// TIA Portal project "Factory_Project_V17" (V17) (continued)
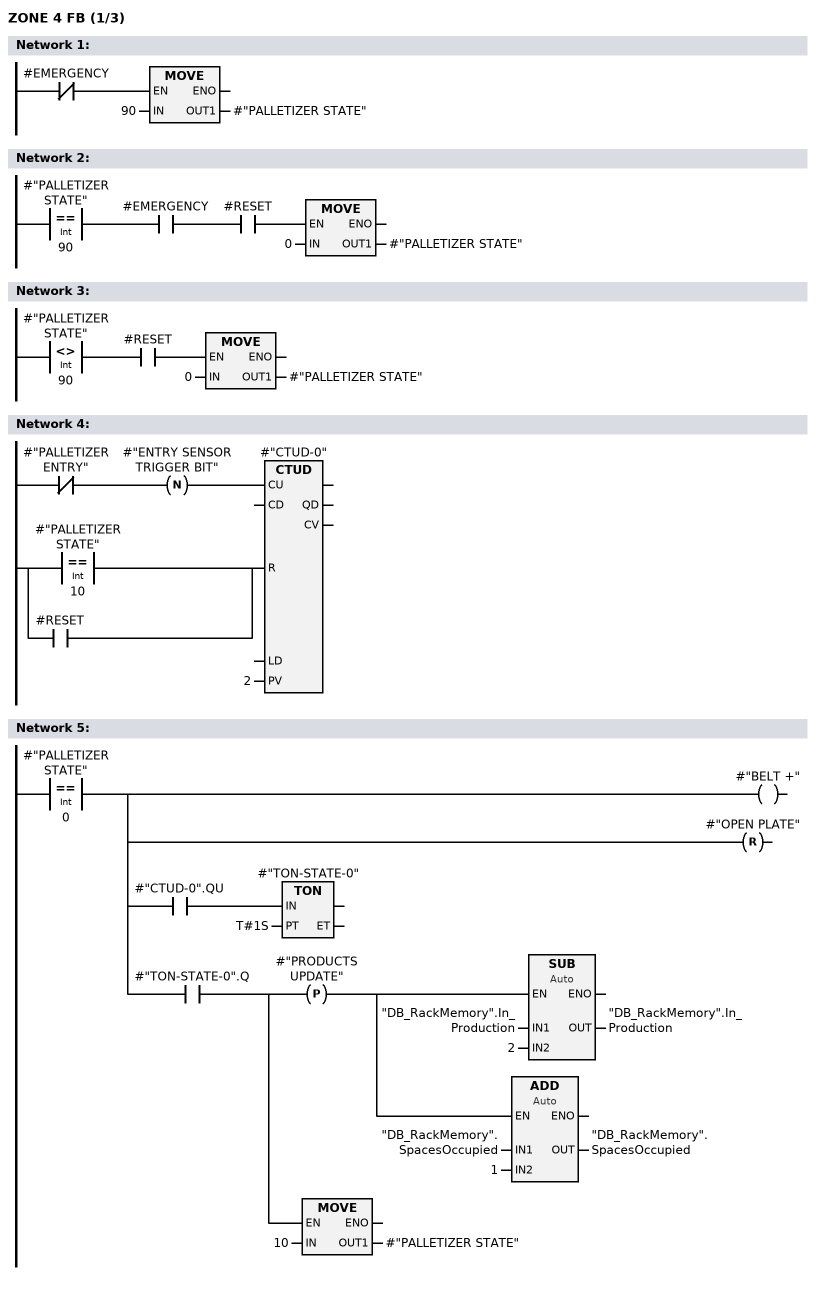
   RUNG wire#powerrail
      I_Contact( #EMERGENCY )
      Move(in := 90, out1 => #"PALLETIZER STATE")
   END_RUNG
   // the same network as SCL:
   IF NOT #EMERGENCY THEN #"PALLETIZER STATE" := 90; END_IF;
END_REGION

REGION Network 2
   RUNG wire#powerrail
      { S7_Templates := "SrcType := Int" } EQ_Contact(in1 := #"PALLETIZER STATE", in2 := 90)
      Contact( #EMERGENCY )
      Contact( #RESET )
      Move(in := 0, out1 => #"PALLETIZER STATE")
   END_RUNG
   // the same network as SCL:
   IF (#"PALLETIZER STATE" = 90) AND #EMERGENCY AND #RESET THEN #"PALLETIZER STATE" := 0; END_IF;
END_REGION

REGION Network 3
   RUNG wire#powerrail
      { S7_Templates := "SrcType := Int" } NE_Contact(in1 := #"PALLETIZER STATE", in2 := 90)
      Contact( #RESET )
      Move(in := 0, out1 => #"PALLETIZER STATE")
   END_RUNG
   // the same network as SCL:
   IF (#"PALLETIZER STATE" <> 90) AND #RESET THEN #"PALLETIZER STATE" := 0; END_IF;
END_REGION

REGION Network 4
   #_w1 := NOT (NOT #"PALLETIZER ENTRY") AND #"ENTRY SENSOR TRIGGER BIT";   // falling edge
   #"ENTRY SENSOR TRIGGER BIT" := NOT #"PALLETIZER ENTRY";
   #"CTUD-0"(CU := #_w1, R := (#"PALLETIZER STATE" = 10) OR #RESET, PV := 2);   // CTUD
END_REGION

REGION Network 5
   #"BELT +" := #"PALLETIZER STATE" = 0;
   IF #"BELT +" THEN #"OPEN PLATE" := FALSE; END_IF;
   #"TON-STATE-0"(IN := #"BELT +" AND #"CTUD-0".QU, PT := T#1S);   // TON
   #_w1 := #"BELT +" AND #"TON-STATE-0".Q;
   #_w2 := #_w1 AND NOT #"PRODUCTS UPDATE";   // rising edge
   #"PRODUCTS UPDATE" := #_w1;
   IF #_w2 THEN
       "DB_RackMemory".In_Production := "DB_RackMemory".In_Production - 2;
       "DB_RackMemory".SpacesOccupied := "DB_RackMemory".SpacesOccupied + 1;
   END_IF;
   IF #_w1 THEN #"PALLETIZER STATE" := 10; END_IF;
END_REGION

REGION Network 6
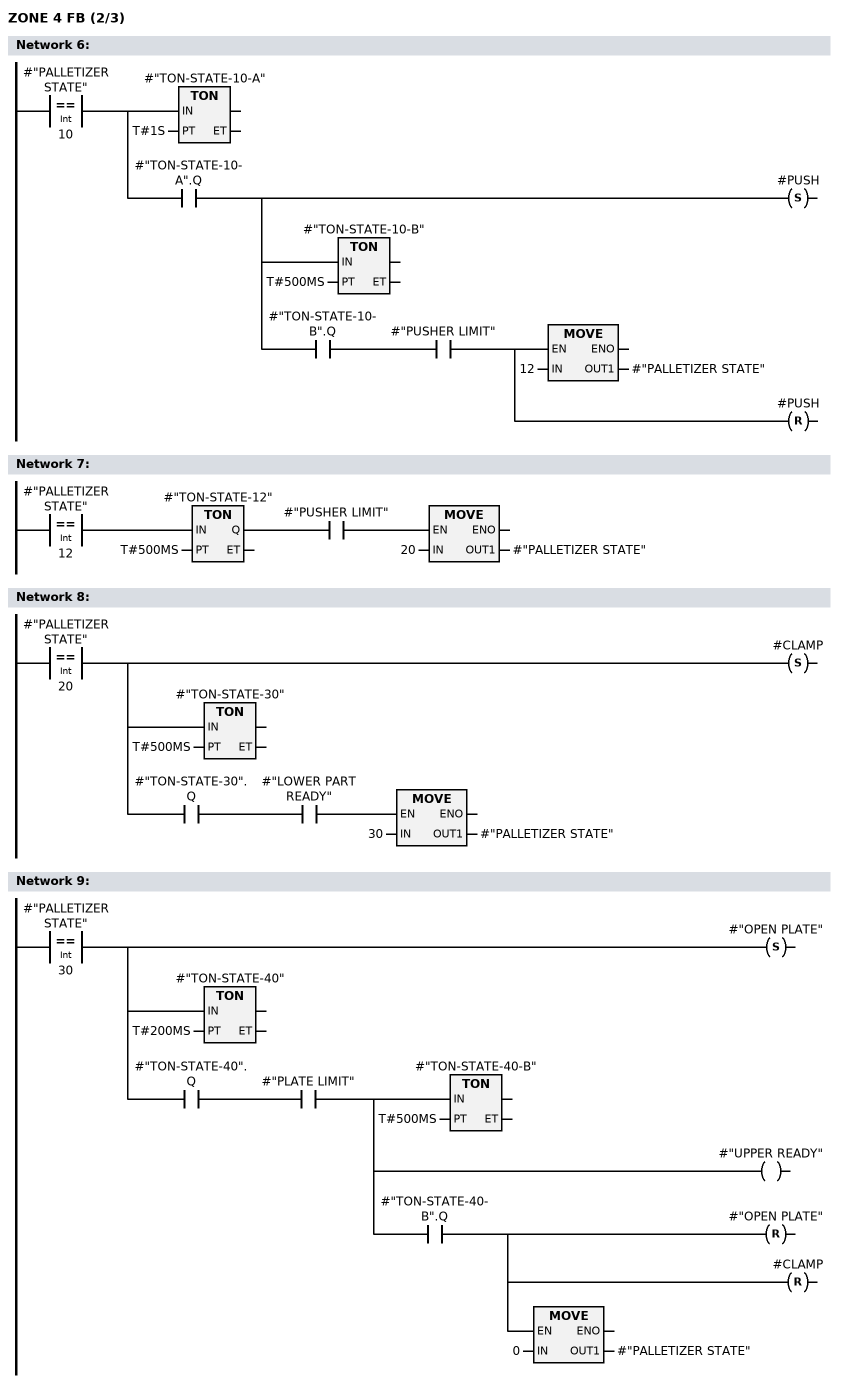
   #_w1 := #"PALLETIZER STATE" = 10;
   #"TON-STATE-10-A"(IN := #_w1, PT := T#1S);   // TON
   #_w2 := #_w1 AND #"TON-STATE-10-A".Q;
   IF #_w2 THEN #PUSH := TRUE; END_IF;
   #"TON-STATE-10-B"(IN := #_w2, PT := T#500MS);   // TON
   IF #_w2 AND #"TON-STATE-10-B".Q AND #"PUSHER LIMIT" THEN
       #"PALLETIZER STATE" := 12;
       #PUSH := FALSE;
   END_IF;
END_REGION

REGION Network 7
   #"TON-STATE-12"(IN := #"PALLETIZER STATE" = 12, PT := T#500MS);   // TON
   IF #"TON-STATE-12".Q AND #"PUSHER LIMIT" THEN #"PALLETIZER STATE" := 20; END_IF;
END_REGION

REGION Network 8
   #_w1 := #"PALLETIZER STATE" = 20;
   IF #_w1 THEN #CLAMP := TRUE; END_IF;
   #"TON-STATE-30"(IN := #_w1, PT := T#500MS);   // TON
   IF #_w1 AND #"TON-STATE-30".Q AND #"LOWER PART READY" THEN #"PALLETIZER STATE" := 30; END_IF;
END_REGION

REGION Network 9
   #_w1 := #"PALLETIZER STATE" = 30;
   IF #_w1 THEN #"OPEN PLATE" := TRUE; END_IF;
   #"TON-STATE-40"(IN := #_w1, PT := T#200MS);   // TON
   #_w2 := #_w1 AND #"TON-STATE-40".Q AND #"PLATE LIMIT";
   #"TON-STATE-40-B"(IN := #_w2, PT := T#500MS);   // TON
   #"UPPER READY" := #_w2;
   IF #_w2 AND #"TON-STATE-40-B".Q THEN
       #"OPEN PLATE" := FALSE;
       #CLAMP := FALSE;
       #"PALLETIZER STATE" := 0;
   END_IF;
END_REGION

REGION Network 10
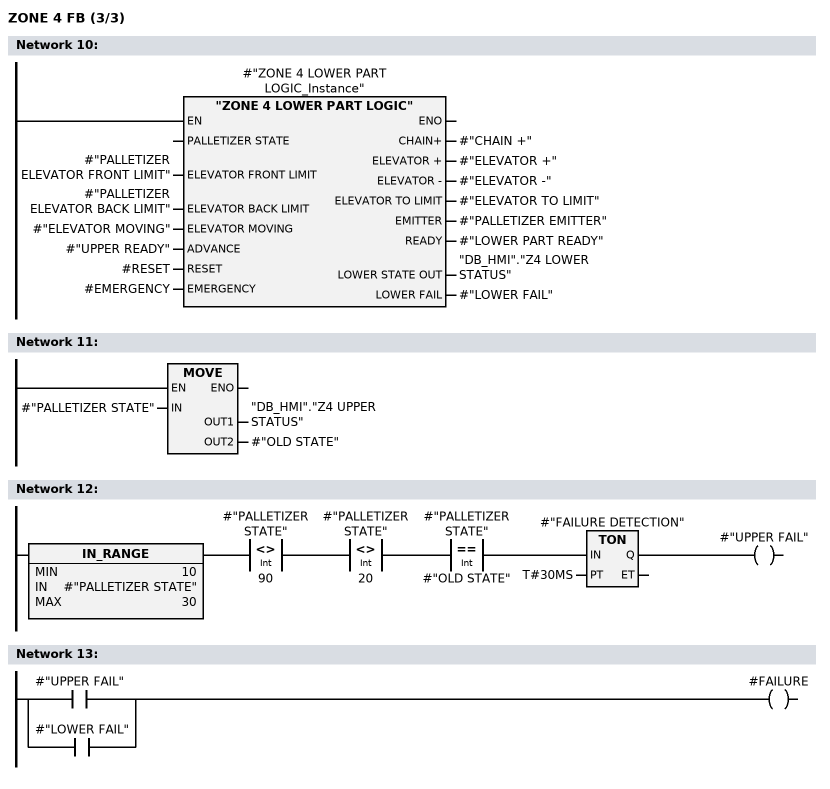
   RUNG wire#powerrail
      #"ZONE 4 LOWER PART LOGIC_Instance"("PALLETIZER STATE" :=, "ELEVATOR FRONT LIMIT" := #"PALLETIZER ELEVATOR FRONT LIMIT", "ELEVATOR BACK LIMIT" := #"PALLETIZER ELEVATOR BACK LIMIT", "ELEVATOR MOVING" := #"ELEVATOR MOVING", ADVANCE := #"UPPER READY", RESET := #RESET, EMERGENCY := #EMERGENCY, "CHAIN+" => #"CHAIN +", "ELEVATOR +" => #"ELEVATOR +", "ELEVATOR -" => #"ELEVATOR -", "ELEVATOR TO LIMIT" => #"ELEVATOR TO LIMIT", EMITTER => #"PALLETIZER EMITTER", READY => #"LOWER PART READY", "LOWER STATE OUT" => "DB_HMI"."Z4 LOWER STATUS", "LOWER FAIL" => #"LOWER FAIL")
   END_RUNG
   // the same network as SCL:
   #"ZONE 4 LOWER PART LOGIC_Instance"("ELEVATOR FRONT LIMIT" := #"PALLETIZER ELEVATOR FRONT LIMIT",   // "ZONE 4 LOWER PART LOGIC"
                           "ELEVATOR BACK LIMIT" := #"PALLETIZER ELEVATOR BACK LIMIT",
                           "ELEVATOR MOVING" := #"ELEVATOR MOVING",
                           ADVANCE := #"UPPER READY",
                           RESET := #RESET,
                           EMERGENCY := #EMERGENCY,
                           "CHAIN+" => #"CHAIN +",
                           "ELEVATOR +" => #"ELEVATOR +",
                           "ELEVATOR -" => #"ELEVATOR -",
                           "ELEVATOR TO LIMIT" => #"ELEVATOR TO LIMIT",
                           EMITTER => #"PALLETIZER EMITTER",
                           READY => #"LOWER PART READY",
                           "LOWER STATE OUT" => "DB_HMI"."Z4 LOWER STATUS",
                           "LOWER FAIL" => #"LOWER FAIL");
END_REGION

REGION Network 11
   RUNG wire#powerrail
      Move(in := #"PALLETIZER STATE", out1 => "DB_HMI"."Z4 UPPER STATUS", out2 => #"OLD STATE")
   END_RUNG
   // the same network as SCL:
   "DB_HMI"."Z4 UPPER STATUS" := #"PALLETIZER STATE";
   #"OLD STATE" := #"PALLETIZER STATE";
END_REGION

REGION Network 12
   #"FAILURE DETECTION"(IN := (10 <= #"PALLETIZER STATE") AND (#"PALLETIZER STATE" <= 30) AND (#"PALLETIZER STATE" <> 90) AND (#"PALLETIZER STATE" <> 20) AND (#"PALLETIZER STATE" = #"OLD STATE"),   // TON
                        PT := T#30MS);
   #"UPPER FAIL" := #"FAILURE DETECTION".Q;
END_REGION

REGION Network 13
   RUNG wire#powerrail
      Contact( #"UPPER FAIL" )
      wire#w1
      Coil( #FAILURE )
   END_RUNG
   RUNG wire#powerrail
      Contact( #"LOWER FAIL" )
   END_RUNG wire#w1
   // the same network as SCL:
   #FAILURE := #"UPPER FAIL" OR #"LOWER FAIL";
END_REGION
END_FUNCTION_BLOCK

FUNCTION_BLOCK "ZONE 4 LOWER PART LOGIC"   // FB17, LAD
{ S7_Optimized_Access := 'TRUE' }
VERSION : 0.1
   VAR_INPUT
      "PALLETIZER STATE" : Int;
      "ELEVATOR FRONT LIMIT" : Bool;
      "ELEVATOR BACK LIMIT" : Bool;
      "ELEVATOR MOVING" : Bool;
      ADVANCE : Bool;
      RESET : Bool;
      EMERGENCY : Bool;
   END_VAR
   VAR_OUTPUT
      "CHAIN+" : Bool;
      "ELEVATOR +" : Bool;
      "ELEVATOR -" : Bool;
      "ELEVATOR TO LIMIT" : Bool;
      EMITTER : Bool;
      READY : Bool;
      "LOWER STATE OUT" : Int;
      "LOWER FAIL" : Bool;
   END_VAR
   VAR
      "LOWER STATE" : Int := 0;
      "TON-ELEVATOR-UP" : TON_TIME;
      "TON-ELEVATOR-DOWN" : TON_TIME;
      "ZONE 4 CHAIN + ELEVATOR_Instance" : "ZONE 4 CHAIN + ELEVATOR";
      "OLD STATE" : Int;
      "FAILURE DETECTION" : TON_TIME;
   END_VAR
   VAR_TEMP   // added for the SCL form of the ladder/FBD networks
      _w1 : Bool;
   END_VAR
BEGIN

REGION Network 1
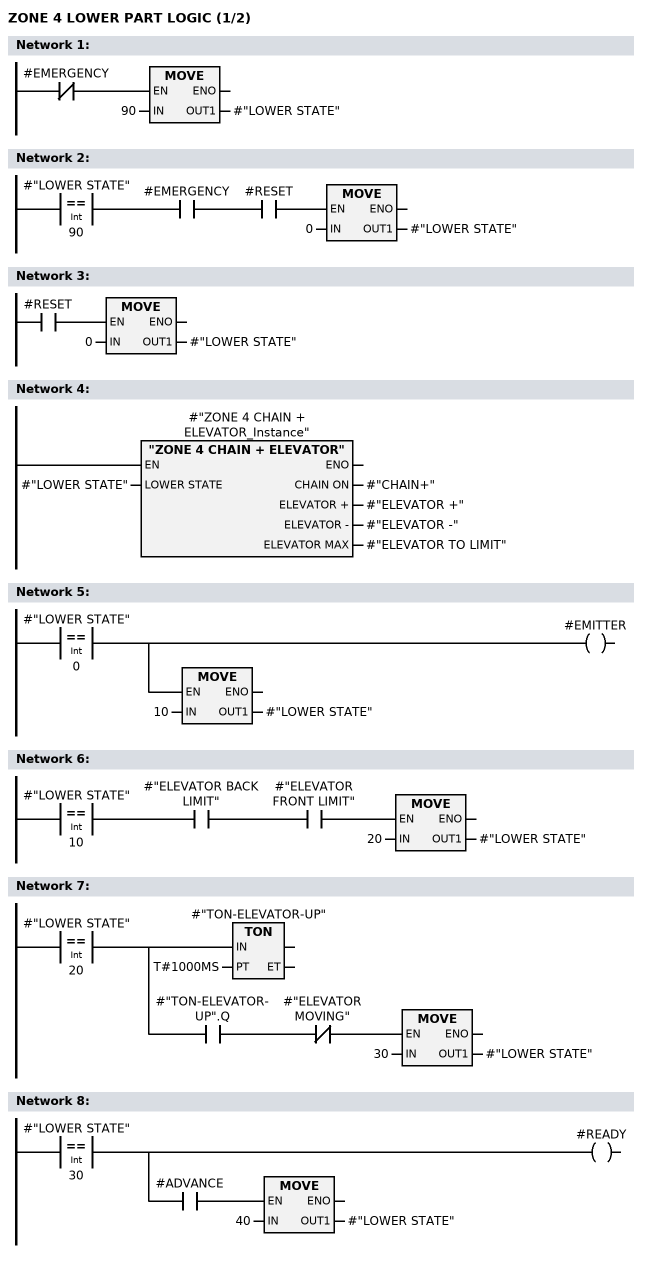
   RUNG wire#powerrail
      I_Contact( #EMERGENCY )
      Move(in := 90, out1 => #"LOWER STATE")
   END_RUNG
   // the same network as SCL:
   IF NOT #EMERGENCY THEN #"LOWER STATE" := 90; END_IF;
END_REGION

REGION Network 2
   RUNG wire#powerrail
      { S7_Templates := "SrcType := Int" } EQ_Contact(in1 := #"LOWER STATE", in2 := 90)
      Contact( #EMERGENCY )
      Contact( #RESET )
      Move(in := 0, out1 => #"LOWER STATE")
   END_RUNG
   // the same network as SCL:
   IF (#"LOWER STATE" = 90) AND #EMERGENCY AND #RESET THEN #"LOWER STATE" := 0; END_IF;
END_REGION

REGION Network 3
   RUNG wire#powerrail
      Contact( #RESET )
      Move(in := 0, out1 => #"LOWER STATE")
   END_RUNG
   // the same network as SCL:
   IF #RESET THEN #"LOWER STATE" := 0; END_IF;
END_REGION

REGION Network 4
   RUNG wire#powerrail
      #"ZONE 4 CHAIN + ELEVATOR_Instance"("LOWER STATE" := #"LOWER STATE", "CHAIN ON" => #"CHAIN+", "ELEVATOR +" => #"ELEVATOR +", "ELEVATOR -" => #"ELEVATOR -", "ELEVATOR MAX" => #"ELEVATOR TO LIMIT")
   END_RUNG
   // the same network as SCL:
   #"ZONE 4 CHAIN + ELEVATOR_Instance"("LOWER STATE" := #"LOWER STATE",   // "ZONE 4 CHAIN + ELEVATOR"
                           "CHAIN ON" => #"CHAIN+",
                           "ELEVATOR +" => #"ELEVATOR +",
                           "ELEVATOR -" => #"ELEVATOR -",
                           "ELEVATOR MAX" => #"ELEVATOR TO LIMIT");
END_REGION

REGION Network 5
   RUNG wire#powerrail
      { S7_Templates := "SrcType := Int" } EQ_Contact(in1 := #"LOWER STATE", in2 := 0)
      wire#w1
      Coil( #EMITTER )
   END_RUNG
   RUNG wire#w1
      Move(in := 10, out1 => #"LOWER STATE")
   END_RUNG
   // the same network as SCL:
   #EMITTER := #"LOWER STATE" = 0;
   IF #EMITTER THEN #"LOWER STATE" := 10; END_IF;
END_REGION

REGION Network 6
   RUNG wire#powerrail
      { S7_Templates := "SrcType := Int" } EQ_Contact(in1 := #"LOWER STATE", in2 := 10)
      Contact( #"ELEVATOR BACK LIMIT" )
      Contact( #"ELEVATOR FRONT LIMIT" )
      Move(in := 20, out1 => #"LOWER STATE")
   END_RUNG
   // the same network as SCL:
   IF (#"LOWER STATE" = 10) AND #"ELEVATOR BACK LIMIT" AND #"ELEVATOR FRONT LIMIT" THEN
       #"LOWER STATE" := 20;
   END_IF;
END_REGION

REGION Network 7
   #_w1 := #"LOWER STATE" = 20;
   #"TON-ELEVATOR-UP"(IN := #_w1, PT := T#1000MS);   // TON
   IF #_w1 AND #"TON-ELEVATOR-UP".Q AND NOT #"ELEVATOR MOVING" THEN #"LOWER STATE" := 30; END_IF;
END_REGION

REGION Network 8
   RUNG wire#powerrail
      { S7_Templates := "SrcType := Int" } EQ_Contact(in1 := #"LOWER STATE", in2 := 30)
      wire#w1
      Coil( #READY )
   END_RUNG
   RUNG wire#w1
      Contact( #ADVANCE )
      Move(in := 40, out1 => #"LOWER STATE")
   END_RUNG
   // the same network as SCL:
   #READY := #"LOWER STATE" = 30;
   IF #READY AND #ADVANCE THEN #"LOWER STATE" := 40; END_IF;
END_REGION

REGION Network 9
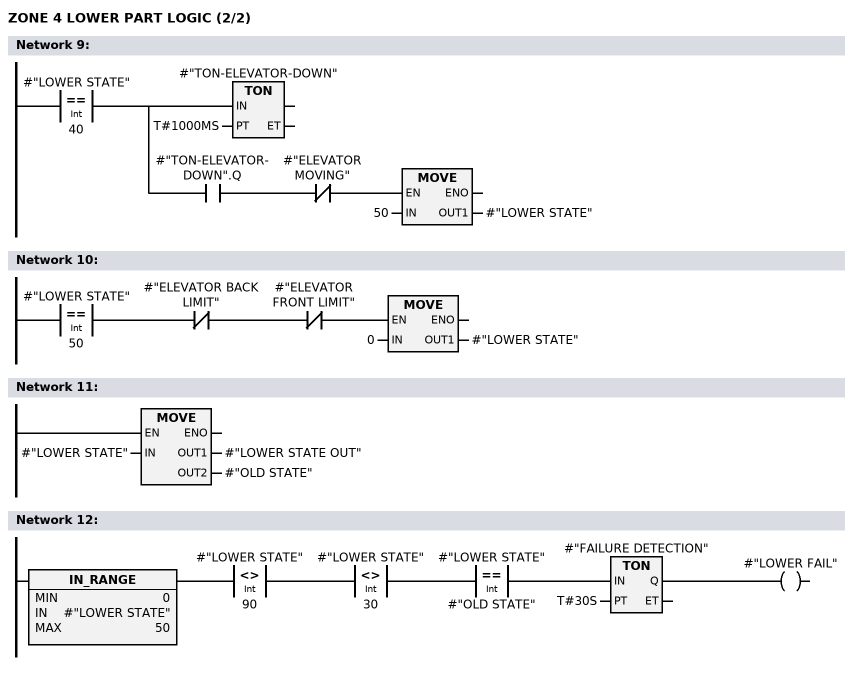
   #_w1 := #"LOWER STATE" = 40;
   #"TON-ELEVATOR-DOWN"(IN := #_w1, PT := T#1000MS);   // TON
   IF #_w1 AND #"TON-ELEVATOR-DOWN".Q AND NOT #"ELEVATOR MOVING" THEN #"LOWER STATE" := 50; END_IF;
END_REGION

REGION Network 10
   RUNG wire#powerrail
      { S7_Templates := "SrcType := Int" } EQ_Contact(in1 := #"LOWER STATE", in2 := 50)
      I_Contact( #"ELEVATOR BACK LIMIT" )
      I_Contact( #"ELEVATOR FRONT LIMIT" )
      Move(in := 0, out1 => #"LOWER STATE")
   END_RUNG
   // the same network as SCL:
   IF (#"LOWER STATE" = 50) AND NOT #"ELEVATOR BACK LIMIT" AND NOT #"ELEVATOR FRONT LIMIT" THEN
       #"LOWER STATE" := 0;
   END_IF;
END_REGION

REGION Network 11
   RUNG wire#powerrail
      Move(in := #"LOWER STATE", out1 => #"LOWER STATE OUT", out2 => #"OLD STATE")
   END_RUNG
   // the same network as SCL:
   #"LOWER STATE OUT" := #"LOWER STATE";
   #"OLD STATE" := #"LOWER STATE";
END_REGION

REGION Network 12
   #"FAILURE DETECTION"(IN := (0 <= #"LOWER STATE") AND (#"LOWER STATE" <= 50) AND (#"LOWER STATE" <> 90) AND (#"LOWER STATE" <> 30) AND (#"LOWER STATE" = #"OLD STATE"),   // TON
                        PT := T#30S);
   #"LOWER FAIL" := #"FAILURE DETECTION".Q;
END_REGION
END_FUNCTION_BLOCK

// folder: ZONE_4_BLOCKS/ZONE 4 SUB BLOCKS

FUNCTION_BLOCK "ZONE 4 CHAIN + ELEVATOR"   // FB18, SCL
{ S7_Optimized_Access := 'TRUE' }
VERSION : 0.1
   VAR_INPUT
      "LOWER STATE" : Int;
   END_VAR
   VAR_OUTPUT
      "CHAIN ON" : Bool;
      "ELEVATOR +" : Bool;
      "ELEVATOR -" : Bool;
      "ELEVATOR MAX" : Bool;
   END_VAR
BEGIN
   CASE #"LOWER STATE" OF
       0:  // Statement section case 1
           #"CHAIN ON":=1;
           #"ELEVATOR +" := 0;
           #"ELEVATOR MAX" := 1;
           #"ELEVATOR -" := 1;
       10:  // Statement section case 2 to 4
           #"CHAIN ON" :=1;
           #"ELEVATOR +" := 0;
           #"ELEVATOR MAX" := 1;
           #"ELEVATOR -" := 1;
       20:
           #"CHAIN ON" := 0;
           #"ELEVATOR +" := 1;
           #"ELEVATOR MAX" := 1;
           #"ELEVATOR -" := 0;
       30:
           #"CHAIN ON" := 0;
           #"ELEVATOR +" := 1;
           #"ELEVATOR MAX" := 1;
           #"ELEVATOR -" := 0;
       40:
           #"CHAIN ON" := 0;
           #"ELEVATOR +" := 0;
           #"ELEVATOR MAX" := 1;
           #"ELEVATOR -" := 1;
       50:
           #"CHAIN ON" := 1;
           #"ELEVATOR +" := 0;
           #"ELEVATOR MAX" := 1;
           #"ELEVATOR -" := 1;
       ELSE  // Statement section ELSE
           #"CHAIN ON" := 0;
           #"ELEVATOR +" := 0;
           #"ELEVATOR MAX" := 0;
           #"ELEVATOR -" := 0;;
   END_CASE;
END_FUNCTION_BLOCK

// folder: Zone _2_Blocks

FUNCTION_BLOCK "Zone_2_FB"   // FB6, LAD
{ S7_Optimized_Access := 'TRUE' }
VERSION : 0.1
   VAR_INPUT
      "entry sensor A" : Bool;
      "entry sensor B" : Bool;
      EMERGENCY : Bool;
      "ERROR A" : Bool;
      "ERROR B" : Bool;
      START : Bool;
      STOP : Bool;
      RESET : Bool;
   END_VAR
   VAR_OUTPUT
      "start A" : Bool;
      "start B" : Bool;
      "Z2 STATE" : Int;
      "A RESET" : Bool;
      "A STOP" : Bool;
      "B RESET" : Bool;
      "B STOP" : Bool;
   END_VAR
   VAR
      STATE : Int;
   END_VAR
   VAR_TEMP   // added for the SCL form of the ladder/FBD networks
      _w1 : Bool;
      _w2 : Bool;
   END_VAR
BEGIN

REGION Network 1
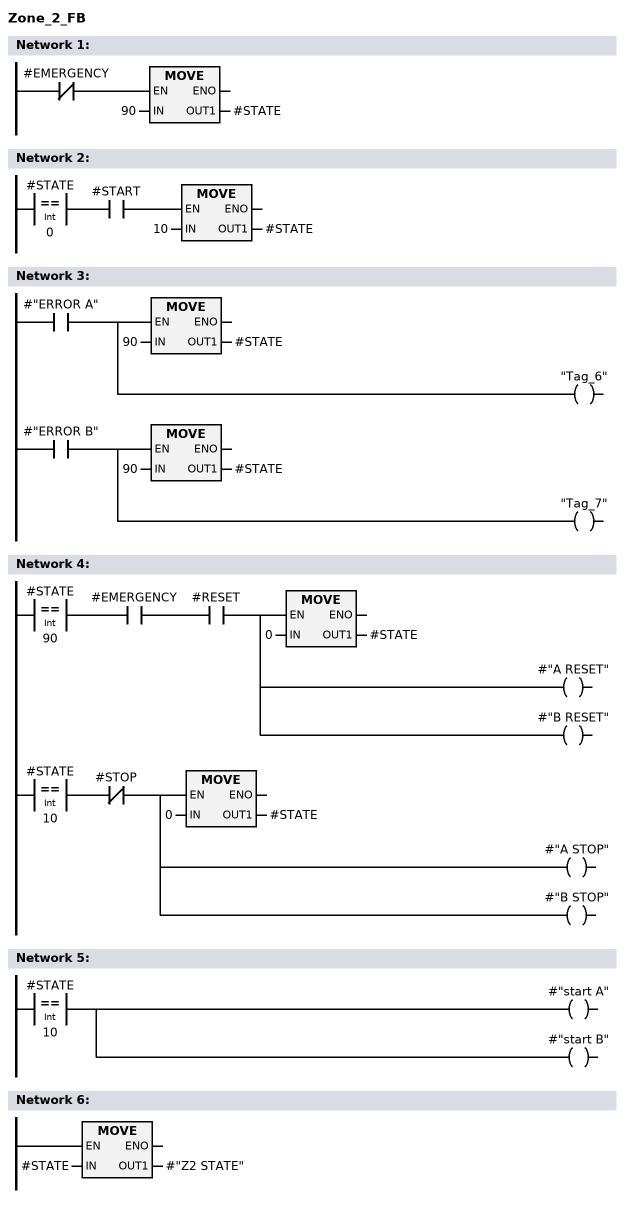
   RUNG wire#powerrail
      I_Contact( #EMERGENCY )
      Move(in := 90, out1 => #STATE)
   END_RUNG
   // the same network as SCL:
   IF NOT #EMERGENCY THEN #STATE := 90; END_IF;
END_REGION

REGION Network 2
   RUNG wire#powerrail
      { S7_Templates := "SrcType := Int" } EQ_Contact(in1 := #STATE, in2 := 0)
      Contact( #START )
      Move(in := 10, out1 => #STATE)
   END_RUNG
   // the same network as SCL:
   IF (#STATE = 0) AND #START THEN #STATE := 10; END_IF;
END_REGION

REGION Network 3
   RUNG wire#powerrail
      Contact( #"ERROR A" )
      wire#w1
      Move(in := 90, out1 => #STATE)
   END_RUNG
   RUNG wire#w1
      Coil( "Tag_6" )
   END_RUNG
   RUNG wire#powerrail
      Contact( #"ERROR B" )
      wire#w2
      Move(in := 90, out1 => #STATE)
   END_RUNG
   RUNG wire#w2
      Coil( "Tag_7" )
   END_RUNG
   // the same network as SCL:
   IF #"ERROR A" THEN #STATE := 90; END_IF;
   "Tag_6" := #"ERROR A";
   IF #"ERROR B" THEN #STATE := 90; END_IF;
   "Tag_7" := #"ERROR B";
END_REGION

REGION Network 4
   RUNG wire#powerrail
      { S7_Templates := "SrcType := Int" } EQ_Contact(in1 := #STATE, in2 := 90)
      Contact( #EMERGENCY )
      Contact( #RESET )
      wire#w1
      Move(in := 0, out1 => #STATE)
   END_RUNG
   RUNG wire#w1
      Coil( #"A RESET" )
   END_RUNG
   RUNG wire#w1
      Coil( #"B RESET" )
   END_RUNG
   RUNG wire#powerrail
      { S7_Templates := "SrcType := Int" } EQ_Contact(in1 := #STATE, in2 := 10)
      I_Contact( #STOP )
      wire#w2
      Move(in := 0, out1 => #STATE)
   END_RUNG
   RUNG wire#w2
      Coil( #"A STOP" )
   END_RUNG
   RUNG wire#w2
      Coil( #"B STOP" )
   END_RUNG
   // the same network as SCL:
   #_w1 := (#STATE = 90) AND #EMERGENCY AND #RESET;
   IF #_w1 THEN #STATE := 0; END_IF;
   #"A RESET" := #_w1;
   #"B RESET" := #_w1;
   #_w2 := (#STATE = 10) AND NOT #STOP;
   IF #_w2 THEN #STATE := 0; END_IF;
   #"A STOP" := #_w2;
   #"B STOP" := #_w2;
END_REGION

REGION Network 5
   RUNG wire#powerrail
      { S7_Templates := "SrcType := Int" } EQ_Contact(in1 := #STATE, in2 := 10)
      wire#w1
      Coil( #"start A" )
   END_RUNG
   RUNG wire#w1
      Coil( #"start B" )
   END_RUNG
   // the same network as SCL:
   #"start A" := #STATE = 10;
   #"start B" := #"start A";
END_REGION

REGION Network 6
   RUNG wire#powerrail
      Move(in := #STATE, out1 => #"Z2 STATE")
   END_RUNG
   // the same network as SCL:
   #"Z2 STATE" := #STATE;
END_REGION
END_FUNCTION_BLOCK

// folder: Zone_3_blocks

FUNCTION_BLOCK "Zone_3_FB"   // FB7, LAD
{ S7_Optimized_Access := 'TRUE' }
VERSION : 0.1
   VAR_INPUT
      START : Bool;
      STOP : Bool;
      EMERGENCY : Bool;
      RESET : Bool;
      "UP ELEVATOR A LEFT SENSOR" : Bool;
      "UP ELEVATOR A RIGHT SENSOR" : Bool;
      "DOWN ELEVATOR A LEFT SENSOR" : Bool;
      "DOWN ELEVATOR A RIGHT SENSOR" : Bool;
      "UP ELEVATOR B LEFT SENSOR" : Bool;
      "UP ELEVATOR B RIGHT SENSOR" : Bool;
      "DOWN ELEVATOR B LEFT SENSOR" : Bool;
      "DOWN ELEVATOR B RIGHT SENSOR" : Bool;
      "BRIDGE A1 SENSOR" : Bool;
      "BRIDGE A2 SENSOR" : Bool;
      "BRIDGE B1 SENSOR" : Bool;
      "BRIDGE B2 SENSOR" : Bool;
      "PRODUCT A AT ASSEMPLY" : Bool;
      "PRODUCT B AT ASSEMPLY" : Bool;
      "PRODUCT LEFT ASSEMPLY" : Bool;
      "POSITIONER A CLAMPED" : Bool;
      "POSITIONER B CLAMPED" : Bool;
      "POSITIONER B LIMIT" : Bool;
      "ASSEMPLER MOVING X" : Bool;
      "ASSEMPLER MOVING Z" : Bool;
      "ASSEMPLER ROATATING" : Bool;
      "ASSEMPLER ITEM DETECTED" : Bool;
      "ASSEMPLER X POSITION" : Real;
      "ASSEMPLER Z POSITION" : Real;
      "UP ELEVATOR A POSITION" : Real;
      "DOWN ELEVATOR A POSITION" : Real;
      "UP ELEVATOR B POSITION" : Real;
      "DOWN ELEVATOR B POSITION" : Real;
      "MACHINE A EXIT SENSOR" : Bool;
      "MACHINE B EXIT SENSOR" : Bool;
   END_VAR
   VAR_OUTPUT
      Z3A1 : Bool;
      Z3A2 : Bool;
      Z3A3 : Bool;
      Z3A4 : Bool;
      Z3A5 : Bool;
      Z3A6 : Bool;
      Z3B1 : Bool;
      Z3B2 : Bool;
      Z3B3 : Bool;
      Z3B4 : Bool;
      Z3B5 : Bool;
      Z3B6 : Bool;
      Z3B7 : Bool;
      "Z3A1 BRIDGE" : Bool;
      "Z3A2 BRIDGE" : Bool;
      "Z3A3 BRIDGE" : Bool;
      "Z3B1 BRIDGE" : Bool;
      "Z3B2 BRIDGE" : Bool;
      "Z3B3 BRIDGE" : Bool;
      "UP ELEVATOR A STOP BLADE" : Bool;
      "DOWN ELEVATOR A STOP BLADE" : Bool;
      "UP ELEVATOR B STOP BLADE" : Bool;
      "DOWN ELEVATOR B STOP BLADE" : Bool;
      "BRIDGE A1 STOP BLADE" : Bool;
      "BRIDGE A2 STOP BLADE" : Bool;
      "BRIDGE B1 STOP BLADE" : Bool;
      "BRIDGE B2 STOP BLADE" : Bool;
      "UP ELEVATOR A SP" : Real;
      "DOWN ELEVATOR A SP" : Real;
      "UP ELEVATOR B SP" : Real;
      "DOWN ELEVATOR B SP" : Real;
      "UP ELEVATOR A +" : Bool;
      "DOWN ELEVATOR A +" : Bool;
      "UP ELEVATOR B +" : Bool;
      "DOWN ELEVATOR B +" : Bool;
      "POSITIONER A CLAMP" : Bool;
      "POSITIONER B CLAMP" : Bool;
      "POSITIONER B RAISE" : Bool;
      "ASSEMPLER X SP" : Real;
      "ASSEMPLER Z SP" : Real;
      "ASSEMPLER GRAB" : Bool;
      "ASSEMPLER ROTATE" : Bool;
      "ASSEMPLER ROT CCW" : Bool;
   END_VAR
   VAR
      "Z3-STATE" : Int;
      "ZONE-3 BUFFER B" : "ZONE-3 BUFFER";
      "ASSEMPLER BUSY" : Bool;
      "BUFFER A READY" : Bool;
      "BUFFER B READY" : Bool;
      "ZONE 3 ASSEMPLER_Instance" : "ZONE 3 ASSEMPLER";
   END_VAR
BEGIN

REGION Network 1
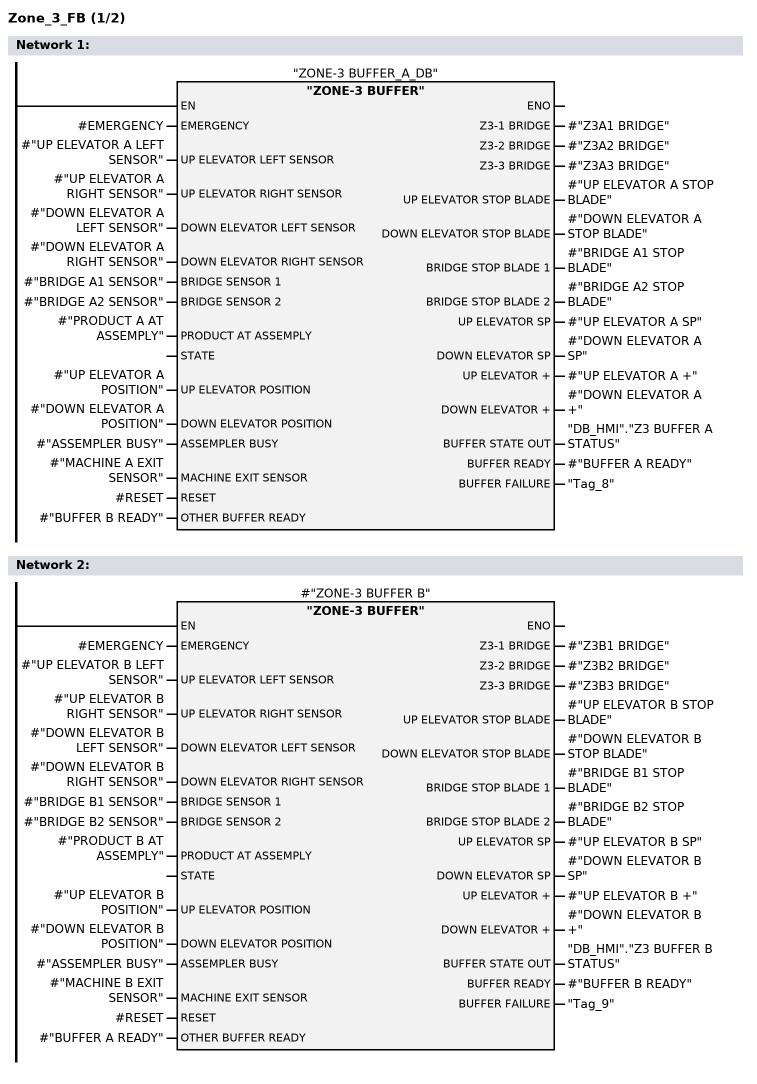
   RUNG wire#powerrail
      "ZONE-3 BUFFER_A_DB"(EMERGENCY := #EMERGENCY, "UP ELEVATOR LEFT SENSOR" := #"UP ELEVATOR A LEFT SENSOR", "UP ELEVATOR RIGHT SENSOR" := #"UP ELEVATOR A RIGHT SENSOR", "DOWN ELEVATOR LEFT SENSOR" := #"DOWN ELEVATOR A LEFT SENSOR", "DOWN ELEVATOR RIGHT SENSOR" := #"DOWN ELEVATOR A RIGHT SENSOR", "BRIDGE SENSOR 1" := #"BRIDGE A1 SENSOR", "BRIDGE SENSOR 2" := #"BRIDGE A2 SENSOR", "PRODUCT AT ASSEMPLY" := #"PRODUCT A AT ASSEMPLY", STATE :=, "UP ELEVATOR POSITION" := #"UP ELEVATOR A POSITION", "DOWN ELEVATOR POSITION" := #"DOWN ELEVATOR A POSITION", "ASSEMPLER BUSY" := #"ASSEMPLER BUSY", "MACHINE EXIT SENSOR" := #"MACHINE A EXIT SENSOR", RESET := #RESET, "OTHER BUFFER READY" := #"BUFFER B READY", "Z3-1 BRIDGE" => #"Z3A1 BRIDGE", "Z3-2 BRIDGE" => #"Z3A2 BRIDGE", "Z3-3 BRIDGE" => #"Z3A3 BRIDGE", "UP ELEVATOR STOP BLADE" => #"UP ELEVATOR A STOP BLADE", "DOWN ELEVATOR STOP BLADE" => #"DOWN ELEVATOR A STOP BLADE", "BRIDGE STOP BLADE 1" => #"BRIDGE A1 STOP BLADE", "BRIDGE STOP BLADE 2" => #"BRIDGE A2 STOP BLADE", "UP ELEVATOR SP" => #"UP ELEVATOR A SP", "DOWN ELEVATOR SP" => #"DOWN ELEVATOR A SP", "UP ELEVATOR +" => #"UP ELEVATOR A +", "DOWN ELEVATOR +" => #"DOWN ELEVATOR A +", "BUFFER STATE OUT" => "DB_HMI"."Z3 BUFFER A STATUS", "BUFFER READY" => #"BUFFER A READY", "BUFFER FAILURE" => "Tag_8")
   END_RUNG
   // the same network as SCL:
   "ZONE-3 BUFFER_A_DB"(EMERGENCY := #EMERGENCY,   // "ZONE-3 BUFFER"
                        "UP ELEVATOR LEFT SENSOR" := #"UP ELEVATOR A LEFT SENSOR",
                        "UP ELEVATOR RIGHT SENSOR" := #"UP ELEVATOR A RIGHT SENSOR",
                        "DOWN ELEVATOR LEFT SENSOR" := #"DOWN ELEVATOR A LEFT SENSOR",
                        "DOWN ELEVATOR RIGHT SENSOR" := #"DOWN ELEVATOR A RIGHT SENSOR",
                        "BRIDGE SENSOR 1" := #"BRIDGE A1 SENSOR",
                        "BRIDGE SENSOR 2" := #"BRIDGE A2 SENSOR",
                        "PRODUCT AT ASSEMPLY" := #"PRODUCT A AT ASSEMPLY",
                        "UP ELEVATOR POSITION" := #"UP ELEVATOR A POSITION",
                        "DOWN ELEVATOR POSITION" := #"DOWN ELEVATOR A POSITION",
                        "ASSEMPLER BUSY" := #"ASSEMPLER BUSY",
                        "MACHINE EXIT SENSOR" := #"MACHINE A EXIT SENSOR",
                        RESET := #RESET,
                        "OTHER BUFFER READY" := #"BUFFER B READY",
                        "Z3-1 BRIDGE" => #"Z3A1 BRIDGE",
                        "Z3-2 BRIDGE" => #"Z3A2 BRIDGE",
                        "Z3-3 BRIDGE" => #"Z3A3 BRIDGE",
                        "UP ELEVATOR STOP BLADE" => #"UP ELEVATOR A STOP BLADE",
                        "DOWN ELEVATOR STOP BLADE" => #"DOWN ELEVATOR A STOP BLADE",
                        "BRIDGE STOP BLADE 1" => #"BRIDGE A1 STOP BLADE",
                        "BRIDGE STOP BLADE 2" => #"BRIDGE A2 STOP BLADE",
                        "UP ELEVATOR SP" => #"UP ELEVATOR A SP",
                        "DOWN ELEVATOR SP" => #"DOWN ELEVATOR A SP",
                        "UP ELEVATOR +" => #"UP ELEVATOR A +",
                        "DOWN ELEVATOR +" => #"DOWN ELEVATOR A +",
                        "BUFFER STATE OUT" => "DB_HMI"."Z3 BUFFER A STATUS",
                        "BUFFER READY" => #"BUFFER A READY",
                        "BUFFER FAILURE" => "Tag_8");
END_REGION

REGION Network 2
   RUNG wire#powerrail
      #"ZONE-3 BUFFER B"(EMERGENCY := #EMERGENCY, "UP ELEVATOR LEFT SENSOR" := #"UP ELEVATOR B LEFT SENSOR", "UP ELEVATOR RIGHT SENSOR" := #"UP ELEVATOR B RIGHT SENSOR", "DOWN ELEVATOR LEFT SENSOR" := #"DOWN ELEVATOR B LEFT SENSOR", "DOWN ELEVATOR RIGHT SENSOR" := #"DOWN ELEVATOR B RIGHT SENSOR", "BRIDGE SENSOR 1" := #"BRIDGE B1 SENSOR", "BRIDGE SENSOR 2" := #"BRIDGE B2 SENSOR", "PRODUCT AT ASSEMPLY" := #"PRODUCT B AT ASSEMPLY", STATE :=, "UP ELEVATOR POSITION" := #"UP ELEVATOR B POSITION", "DOWN ELEVATOR POSITION" := #"DOWN ELEVATOR B POSITION", "ASSEMPLER BUSY" := #"ASSEMPLER BUSY", "MACHINE EXIT SENSOR" := #"MACHINE B EXIT SENSOR", RESET := #RESET, "OTHER BUFFER READY" := #"BUFFER A READY", "Z3-1 BRIDGE" => #"Z3B1 BRIDGE", "Z3-2 BRIDGE" => #"Z3B2 BRIDGE", "Z3-3 BRIDGE" => #"Z3B3 BRIDGE", "UP ELEVATOR STOP BLADE" => #"UP ELEVATOR B STOP BLADE", "DOWN ELEVATOR STOP BLADE" => #"DOWN ELEVATOR B STOP BLADE", "BRIDGE STOP BLADE 1" => #"BRIDGE B1 STOP BLADE", "BRIDGE STOP BLADE 2" => #"BRIDGE B2 STOP BLADE", "UP ELEVATOR SP" => #"UP ELEVATOR B SP", "DOWN ELEVATOR SP" => #"DOWN ELEVATOR B SP", "UP ELEVATOR +" => #"UP ELEVATOR B +", "DOWN ELEVATOR +" => #"DOWN ELEVATOR B +", "BUFFER STATE OUT" => "DB_HMI"."Z3 BUFFER B STATUS", "BUFFER READY" => #"BUFFER B READY", "BUFFER FAILURE" => "Tag_9")
   END_RUNG
   // the same network as SCL:
   #"ZONE-3 BUFFER B"(EMERGENCY := #EMERGENCY,   // "ZONE-3 BUFFER"
                      "UP ELEVATOR LEFT SENSOR" := #"UP ELEVATOR B LEFT SENSOR",
                      "UP ELEVATOR RIGHT SENSOR" := #"UP ELEVATOR B RIGHT SENSOR",
                      "DOWN ELEVATOR LEFT SENSOR" := #"DOWN ELEVATOR B LEFT SENSOR",
                      "DOWN ELEVATOR RIGHT SENSOR" := #"DOWN ELEVATOR B RIGHT SENSOR",
                      "BRIDGE SENSOR 1" := #"BRIDGE B1 SENSOR",
                      "BRIDGE SENSOR 2" := #"BRIDGE B2 SENSOR",
                      "PRODUCT AT ASSEMPLY" := #"PRODUCT B AT ASSEMPLY",
                      "UP ELEVATOR POSITION" := #"UP ELEVATOR B POSITION",
                      "DOWN ELEVATOR POSITION" := #"DOWN ELEVATOR B POSITION",
                      "ASSEMPLER BUSY" := #"ASSEMPLER BUSY",
                      "MACHINE EXIT SENSOR" := #"MACHINE B EXIT SENSOR",
                      RESET := #RESET,
                      "OTHER BUFFER READY" := #"BUFFER A READY",
                      "Z3-1 BRIDGE" => #"Z3B1 BRIDGE",
                      "Z3-2 BRIDGE" => #"Z3B2 BRIDGE",
                      "Z3-3 BRIDGE" => #"Z3B3 BRIDGE",
                      "UP ELEVATOR STOP BLADE" => #"UP ELEVATOR B STOP BLADE",
                      "DOWN ELEVATOR STOP BLADE" => #"DOWN ELEVATOR B STOP BLADE",
                      "BRIDGE STOP BLADE 1" => #"BRIDGE B1 STOP BLADE",
                      "BRIDGE STOP BLADE 2" => #"BRIDGE B2 STOP BLADE",
                      "UP ELEVATOR SP" => #"UP ELEVATOR B SP",
                      "DOWN ELEVATOR SP" => #"DOWN ELEVATOR B SP",
                      "UP ELEVATOR +" => #"UP ELEVATOR B +",
                      "DOWN ELEVATOR +" => #"DOWN ELEVATOR B +",
                      "BUFFER STATE OUT" => "DB_HMI"."Z3 BUFFER B STATUS",
                      "BUFFER READY" => #"BUFFER B READY",
                      "BUFFER FAILURE" => "Tag_9");
END_REGION

REGION Network 3
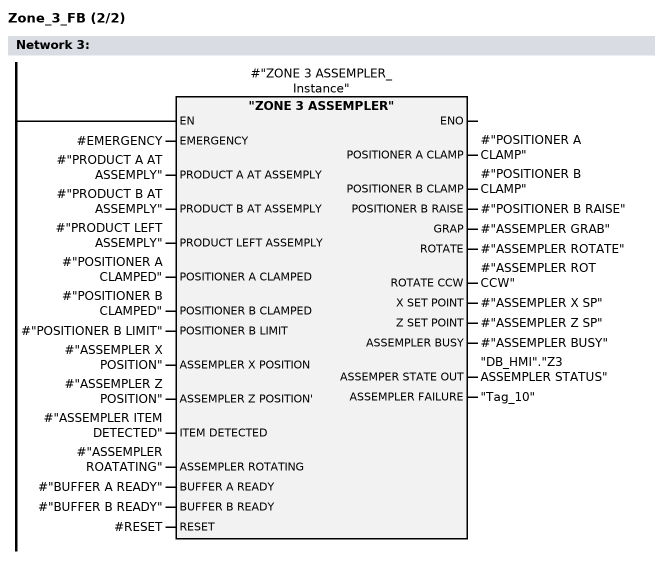
   RUNG wire#powerrail
      #"ZONE 3 ASSEMPLER_Instance"(EMERGENCY := #EMERGENCY, "PRODUCT A AT ASSEMPLY" := #"PRODUCT A AT ASSEMPLY", "PRODUCT B AT ASSEMPLY" := #"PRODUCT B AT ASSEMPLY", "PRODUCT LEFT ASSEMPLY" := #"PRODUCT LEFT ASSEMPLY", "POSITIONER A CLAMPED" := #"POSITIONER A CLAMPED", "POSITIONER B CLAMPED" := #"POSITIONER B CLAMPED", "POSITIONER B LIMIT" := #"POSITIONER B LIMIT", "ASSEMPLER X POSITION" := #"ASSEMPLER X POSITION", "ASSEMPLER Z POSITION'" := #"ASSEMPLER Z POSITION", "ITEM DETECTED" := #"ASSEMPLER ITEM DETECTED", "ASSEMPLER ROTATING" := #"ASSEMPLER ROATATING", "BUFFER A READY" := #"BUFFER A READY", "BUFFER B READY" := #"BUFFER B READY", RESET := #RESET, "POSITIONER A CLAMP" => #"POSITIONER A CLAMP", "POSITIONER B CLAMP" => #"POSITIONER B CLAMP", "POSITIONER B RAISE" => #"POSITIONER B RAISE", GRAP => #"ASSEMPLER GRAB", ROTATE => #"ASSEMPLER ROTATE", "ROTATE CCW" => #"ASSEMPLER ROT CCW", "X SET POINT" => #"ASSEMPLER X SP", "Z SET POINT" => #"ASSEMPLER Z SP", "ASSEMPLER BUSY" => #"ASSEMPLER BUSY", "ASSEMPER STATE OUT" => "DB_HMI"."Z3 ASSEMPLER STATUS", "ASSEMPLER FAILURE" => "Tag_10")
   END_RUNG
   // the same network as SCL:
   #"ZONE 3 ASSEMPLER_Instance"(EMERGENCY := #EMERGENCY,   // "ZONE 3 ASSEMPLER"
                           "PRODUCT A AT ASSEMPLY" := #"PRODUCT A AT ASSEMPLY",
                           "PRODUCT B AT ASSEMPLY" := #"PRODUCT B AT ASSEMPLY",
                           "PRODUCT LEFT ASSEMPLY" := #"PRODUCT LEFT ASSEMPLY",
                           "POSITIONER A CLAMPED" := #"POSITIONER A CLAMPED",
                           "POSITIONER B CLAMPED" := #"POSITIONER B CLAMPED",
                           "POSITIONER B LIMIT" := #"POSITIONER B LIMIT",
                           "ASSEMPLER X POSITION" := #"ASSEMPLER X POSITION",
                           "ASSEMPLER Z POSITION'" := #"ASSEMPLER Z POSITION",
                           "ITEM DETECTED" := #"ASSEMPLER ITEM DETECTED",
                           "ASSEMPLER ROTATING" := #"ASSEMPLER ROATATING",
                           "BUFFER A READY" := #"BUFFER A READY",
                           "BUFFER B READY" := #"BUFFER B READY",
                           RESET := #RESET,
                           "POSITIONER A CLAMP" => #"POSITIONER A CLAMP",
                           "POSITIONER B CLAMP" => #"POSITIONER B CLAMP",
                           "POSITIONER B RAISE" => #"POSITIONER B RAISE",
                           GRAP => #"ASSEMPLER GRAB",
                           ROTATE => #"ASSEMPLER ROTATE",
                           "ROTATE CCW" => #"ASSEMPLER ROT CCW",
                           "X SET POINT" => #"ASSEMPLER X SP",
                           "Z SET POINT" => #"ASSEMPLER Z SP",
                           "ASSEMPLER BUSY" => #"ASSEMPLER BUSY",
                           "ASSEMPER STATE OUT" => "DB_HMI"."Z3 ASSEMPLER STATUS",
                           "ASSEMPLER FAILURE" => "Tag_10");
END_REGION
END_FUNCTION_BLOCK

FUNCTION_BLOCK "ZONE-3 BUFFER"   // FB8, LAD
{ S7_Optimized_Access := 'TRUE' }
VERSION : 0.1
   VAR_INPUT
      EMERGENCY : Bool;
      "UP ELEVATOR LEFT SENSOR" : Bool;
      "UP ELEVATOR RIGHT SENSOR" : Bool;
      "DOWN ELEVATOR LEFT SENSOR" : Bool;
      "DOWN ELEVATOR RIGHT SENSOR" : Bool;
      "BRIDGE SENSOR 1" : Bool;
      "BRIDGE SENSOR 2" : Bool;
      "PRODUCT AT ASSEMPLY" : Bool;
      STATE : Int;
      "UP ELEVATOR POSITION" : Real;
      "DOWN ELEVATOR POSITION" : Real;
      "ASSEMPLER BUSY" : Bool;
      "MACHINE EXIT SENSOR" : Bool;
      RESET : Bool;
      "OTHER BUFFER READY" : Bool;
   END_VAR
   VAR_OUTPUT
      "Z3-1 BRIDGE" : Bool;
      "Z3-2 BRIDGE" : Bool;
      "Z3-3 BRIDGE" : Bool;
      "UP ELEVATOR STOP BLADE" : Bool;
      "DOWN ELEVATOR STOP BLADE" : Bool;
      "BRIDGE STOP BLADE 1" : Bool;
      "BRIDGE STOP BLADE 2" : Bool;
      "UP ELEVATOR SP" : Real;
      "DOWN ELEVATOR SP" : Real;
      "UP ELEVATOR +" : Bool;
      "DOWN ELEVATOR +" : Bool;
      "BUFFER STATE OUT" : Int;
      "BUFFER READY" : Bool;
      "BUFFER FAILURE" : Bool;
   END_VAR
   VAR
      "BUFFER STATE" : Int := 0;
      "OLD BUFFER STATE" : Int;
      "UP ELEVATOR N TRIG LEFT" : Bool;
   END_VAR
   VAR RETAIN
      BUFFER_ITEMS_COUNT : CTUD_INT;
   END_VAR
   VAR
      "DOWN ELEVATOR N TRIG LEFT" : Bool;
      "UP ELEVATOR N TRIG RIGHT" : Bool;
      "BRIDGE SENSOR 2 N TRIG STATE 30" : Bool;
      "BRIDGE SENSOR 1 N TRIG STATE 30" : Bool;
      "ZONE 3 STOP BLADES LOGIC_Instance" : "ZONE 3 STOP BLADES LOGIC";
      "DOWN ELEVATOR RIGHT SENSOR N TRIG" : Bool;
      "ZONE 3 ADVANCING THE BUFFER_Instance" : "ZONE 3 ADVANCING THE BUFFER";
      "ZONE 3 ELEVATORS LOGIC_Instance" : "ZONE 3 ELEVATORS LOGIC";
      "ZONE 3 BRIDGE CONVS LOGIC_Instance" : "ZONE 3 BRIDGE CONVS LOGIC";
      "STATE 30 DONE" : Bool;
      "STATE 50 DONE" : Bool;
      "up right n trig 2" : Bool;
      "down left n trig 2" : Bool;
      processing : Bool;
      "FAILURE DETECTION" : TON_TIME;
   END_VAR
   VAR_TEMP   // added for the SCL form of the ladder/FBD networks
      _w1 : Bool;
      _w2 : Bool;
      _w3 : Bool;
      _w4 : Bool;
   END_VAR
BEGIN

REGION Network 1
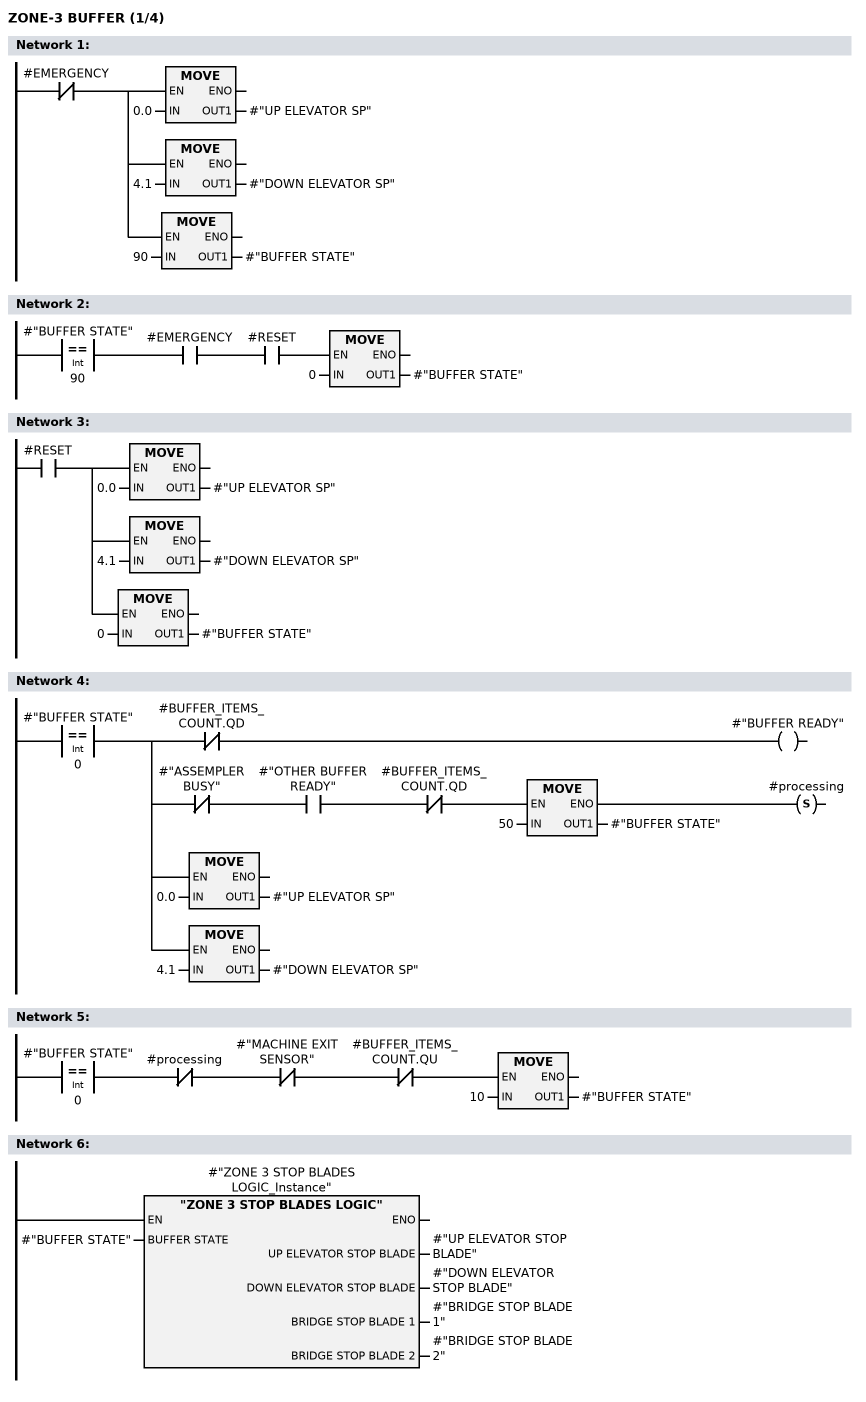
   RUNG wire#powerrail
      I_Contact( #EMERGENCY )
      wire#w1
      Move(in := 0.0, out1 => #"UP ELEVATOR SP")
   END_RUNG
   RUNG wire#w1
      Move(in := 4.1, out1 => #"DOWN ELEVATOR SP")
   END_RUNG
   RUNG wire#w1
      Move(in := 90, out1 => #"BUFFER STATE")
   END_RUNG
   // the same network as SCL:
   IF NOT #EMERGENCY THEN
       #"UP ELEVATOR SP" := 0.0;
       #"DOWN ELEVATOR SP" := 4.1;
       #"BUFFER STATE" := 90;
   END_IF;
END_REGION

REGION Network 2
   RUNG wire#powerrail
      { S7_Templates := "SrcType := Int" } EQ_Contact(in1 := #"BUFFER STATE", in2 := 90)
      Contact( #EMERGENCY )
      Contact( #RESET )
      Move(in := 0, out1 => #"BUFFER STATE")
   END_RUNG
   // the same network as SCL:
   IF (#"BUFFER STATE" = 90) AND #EMERGENCY AND #RESET THEN #"BUFFER STATE" := 0; END_IF;
END_REGION

REGION Network 3
   RUNG wire#powerrail
      Contact( #RESET )
      wire#w1
      Move(in := 0.0, out1 => #"UP ELEVATOR SP")
   END_RUNG
   RUNG wire#w1
      Move(in := 4.1, out1 => #"DOWN ELEVATOR SP")
   END_RUNG
   RUNG wire#w1
      Move(in := 0, out1 => #"BUFFER STATE")
   END_RUNG
   // the same network as SCL:
   IF #RESET THEN
       #"UP ELEVATOR SP" := 0.0;
       #"DOWN ELEVATOR SP" := 4.1;
       #"BUFFER STATE" := 0;
   END_IF;
END_REGION

REGION Network 4
   RUNG wire#powerrail
      { S7_Templates := "SrcType := Int" } EQ_Contact(in1 := #"BUFFER STATE", in2 := 0)
      wire#w1
      I_Contact( #BUFFER_ITEMS_COUNT.QD )
      Coil( #"BUFFER READY" )
   END_RUNG
   RUNG wire#w1
      I_Contact( #"ASSEMPLER BUSY" )
      Contact( #"OTHER BUFFER READY" )
      I_Contact( #BUFFER_ITEMS_COUNT.QD )
      Move(in := 50, out1 => #"BUFFER STATE")
      S_Coil( #processing )
   END_RUNG
   RUNG wire#w1
      Move(in := 0.0, out1 => #"UP ELEVATOR SP")
   END_RUNG
   RUNG wire#w1
      Move(in := 4.1, out1 => #"DOWN ELEVATOR SP")
   END_RUNG
   // the same network as SCL:
   #_w1 := #"BUFFER STATE" = 0;
   #"BUFFER READY" := #_w1 AND NOT #BUFFER_ITEMS_COUNT.QD;
   IF #_w1 AND NOT #"ASSEMPLER BUSY" AND #"OTHER BUFFER READY" AND NOT #BUFFER_ITEMS_COUNT.QD THEN
       #"BUFFER STATE" := 50;
       #processing := TRUE;
   END_IF;
   IF #_w1 THEN
       #"UP ELEVATOR SP" := 0.0;
       #"DOWN ELEVATOR SP" := 4.1;
   END_IF;
END_REGION

